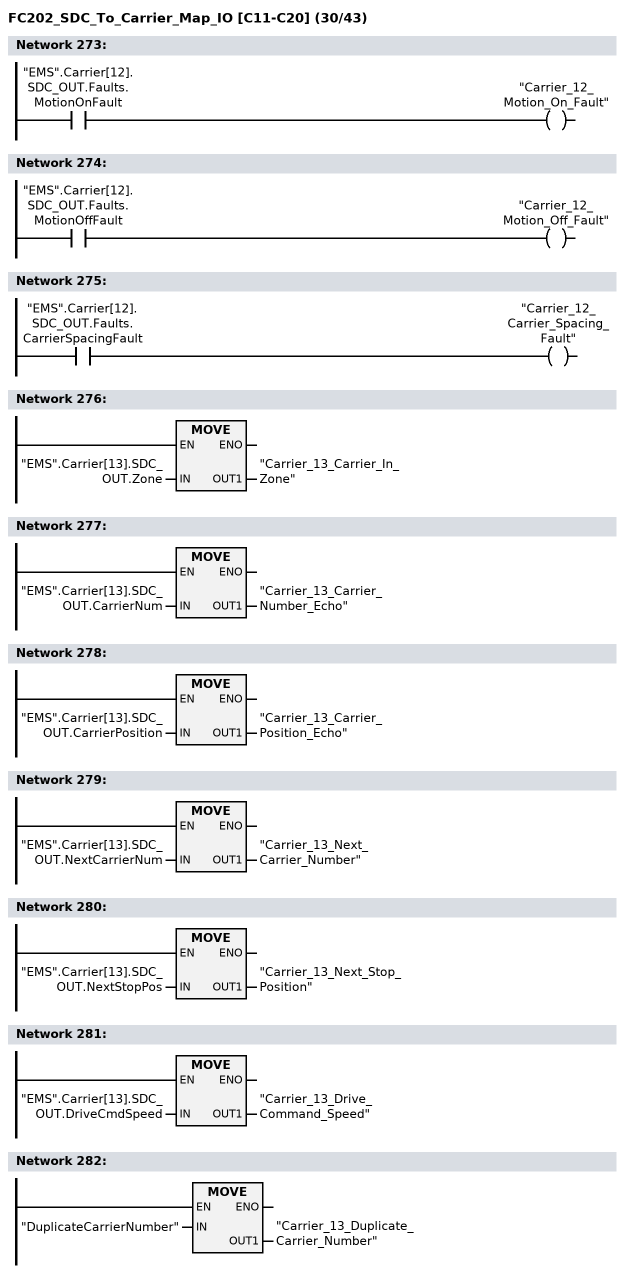
   RUNG wire#powerrail
      Contact( "EMS".Carrier[12].SDC_OUT.Faults.MotionOnFault )
      Coil( "Carrier_12_Motion_On_Fault" )
   END_RUNG
   // the same network as SCL:
   "Carrier_12_Motion_On_Fault" := "EMS".Carrier[12].SDC_OUT.Faults.MotionOnFault;
END_REGION

REGION Network 274
   RUNG wire#powerrail
      Contact( "EMS".Carrier[12].SDC_OUT.Faults.MotionOffFault )
      Coil( "Carrier_12_Motion_Off_Fault" )
   END_RUNG
   // the same network as SCL:
   "Carrier_12_Motion_Off_Fault" := "EMS".Carrier[12].SDC_OUT.Faults.MotionOffFault;
END_REGION

REGION Network 275
   RUNG wire#powerrail
      Contact( "EMS".Carrier[12].SDC_OUT.Faults.CarrierSpacingFault )
      Coil( "Carrier_12_Carrier_Spacing_Fault" )
   END_RUNG
   // the same network as SCL:
   "Carrier_12_Carrier_Spacing_Fault" := "EMS".Carrier[12].SDC_OUT.Faults.CarrierSpacingFault;
END_REGION

REGION Network 276
   RUNG wire#powerrail
      Move(in := "EMS".Carrier[13].SDC_OUT.Zone, out1 => "Carrier_13_Carrier_In_Zone")
   END_RUNG
   // the same network as SCL:
   "Carrier_13_Carrier_In_Zone" := "EMS".Carrier[13].SDC_OUT.Zone;
END_REGION

REGION Network 277
   RUNG wire#powerrail
      Move(in := "EMS".Carrier[13].SDC_OUT.CarrierNum, out1 => "Carrier_13_Carrier_Number_Echo")
   END_RUNG
   // the same network as SCL:
   "Carrier_13_Carrier_Number_Echo" := "EMS".Carrier[13].SDC_OUT.CarrierNum;
END_REGION

REGION Network 278
   RUNG wire#powerrail
      Move(in := "EMS".Carrier[13].SDC_OUT.CarrierPosition, out1 => "Carrier_13_Carrier_Position_Echo")
   END_RUNG
   // the same network as SCL:
   "Carrier_13_Carrier_Position_Echo" := "EMS".Carrier[13].SDC_OUT.CarrierPosition;
END_REGION

REGION Network 279
   RUNG wire#powerrail
      Move(in := "EMS".Carrier[13].SDC_OUT.NextCarrierNum, out1 => "Carrier_13_Next_Carrier_Number")
   END_RUNG
   // the same network as SCL:
   "Carrier_13_Next_Carrier_Number" := "EMS".Carrier[13].SDC_OUT.NextCarrierNum;
END_REGION

REGION Network 280
   RUNG wire#powerrail
      Move(in := "EMS".Carrier[13].SDC_OUT.NextStopPos, out1 => "Carrier_13_Next_Stop_Position")
   END_RUNG
   // the same network as SCL:
   "Carrier_13_Next_Stop_Position" := "EMS".Carrier[13].SDC_OUT.NextStopPos;
END_REGION

REGION Network 281
   RUNG wire#powerrail
      Move(in := "EMS".Carrier[13].SDC_OUT.DriveCmdSpeed, out1 => "Carrier_13_Drive_Command_Speed")
   END_RUNG
   // the same network as SCL:
   "Carrier_13_Drive_Command_Speed" := "EMS".Carrier[13].SDC_OUT.DriveCmdSpeed;
END_REGION

REGION Network 282
   RUNG wire#powerrail
      Move(in := "DuplicateCarrierNumber", out1 => "Carrier_13_Duplicate_Carrier_Number")
   END_RUNG
   // the same network as SCL:
   "Carrier_13_Duplicate_Carrier_Number" := "DuplicateCarrierNumber";
END_REGION

REGION Network 283
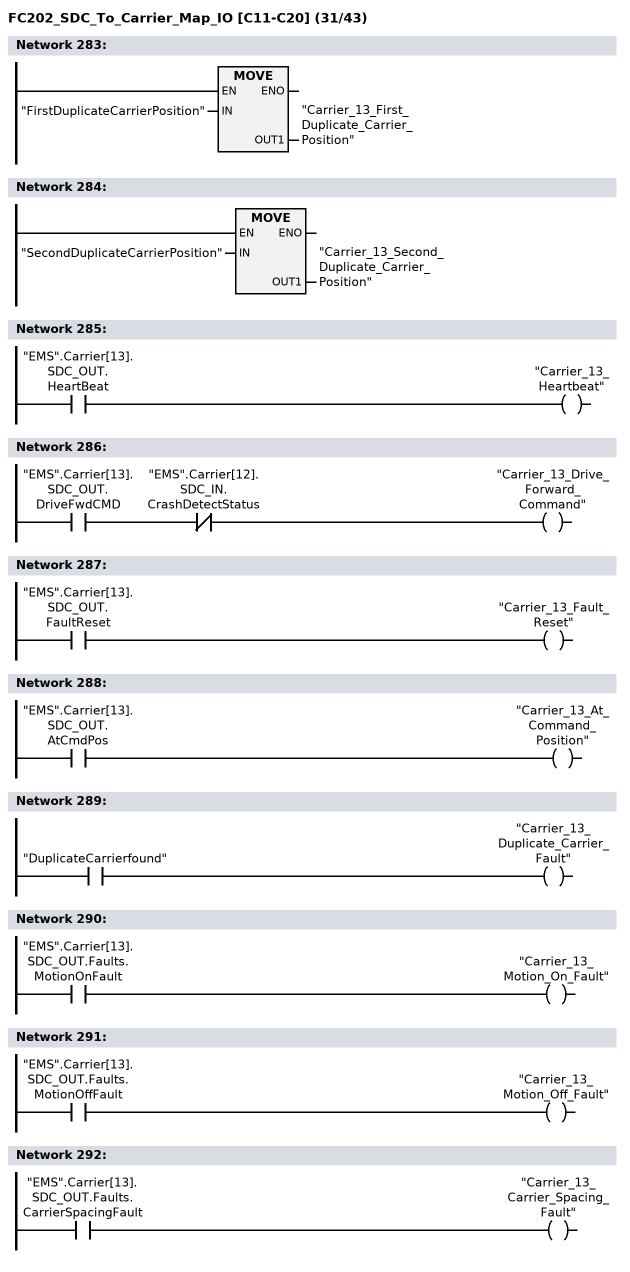
   RUNG wire#powerrail
      Move(in := "FirstDuplicateCarrierPosition", out1 => "Carrier_13_First_Duplicate_Carrier_Position")
   END_RUNG
   // the same network as SCL:
   "Carrier_13_First_Duplicate_Carrier_Position" := "FirstDuplicateCarrierPosition";
END_REGION

REGION Network 284
   RUNG wire#powerrail
      Move(in := "SecondDuplicateCarrierPosition", out1 => "Carrier_13_Second_Duplicate_Carrier_Position")
   END_RUNG
   // the same network as SCL:
   "Carrier_13_Second_Duplicate_Carrier_Position" := "SecondDuplicateCarrierPosition";
END_REGION

REGION Network 285
   RUNG wire#powerrail
      Contact( "EMS".Carrier[13].SDC_OUT.HeartBeat )
      Coil( "Carrier_13_Heartbeat" )
   END_RUNG
   // the same network as SCL:
   "Carrier_13_Heartbeat" := "EMS".Carrier[13].SDC_OUT.HeartBeat;
END_REGION

REGION Network 286
   RUNG wire#powerrail
      Contact( "EMS".Carrier[13].SDC_OUT.DriveFwdCMD )
      I_Contact( "EMS".Carrier[12].SDC_IN.CrashDetectStatus )
      Coil( "Carrier_13_Drive_Forward_Command" )
   END_RUNG
   // the same network as SCL:
   "Carrier_13_Drive_Forward_Command" := "EMS".Carrier[13].SDC_OUT.DriveFwdCMD AND NOT "EMS".Carrier[12].SDC_IN.CrashDetectStatus;
END_REGION

REGION Network 287
   RUNG wire#powerrail
      Contact( "EMS".Carrier[13].SDC_OUT.FaultReset )
      Coil( "Carrier_13_Fault_Reset" )
   END_RUNG
   // the same network as SCL:
   "Carrier_13_Fault_Reset" := "EMS".Carrier[13].SDC_OUT.FaultReset;
END_REGION

REGION Network 288
   RUNG wire#powerrail
      Contact( "EMS".Carrier[13].SDC_OUT.AtCmdPos )
      Coil( "Carrier_13_At_Command_Position" )
   END_RUNG
   // the same network as SCL:
   "Carrier_13_At_Command_Position" := "EMS".Carrier[13].SDC_OUT.AtCmdPos;
END_REGION

REGION Network 289
   RUNG wire#powerrail
      Contact( "DuplicateCarrierfound" )
      Coil( "Carrier_13_Duplicate_Carrier_Fault" )
   END_RUNG
   // the same network as SCL:
   "Carrier_13_Duplicate_Carrier_Fault" := "DuplicateCarrierfound";
END_REGION

REGION Network 290
   RUNG wire#powerrail
      Contact( "EMS".Carrier[13].SDC_OUT.Faults.MotionOnFault )
      Coil( "Carrier_13_Motion_On_Fault" )
   END_RUNG
   // the same network as SCL:
   "Carrier_13_Motion_On_Fault" := "EMS".Carrier[13].SDC_OUT.Faults.MotionOnFault;
END_REGION

REGION Network 291
   RUNG wire#powerrail
      Contact( "EMS".Carrier[13].SDC_OUT.Faults.MotionOffFault )
      Coil( "Carrier_13_Motion_Off_Fault" )
   END_RUNG
   // the same network as SCL:
   "Carrier_13_Motion_Off_Fault" := "EMS".Carrier[13].SDC_OUT.Faults.MotionOffFault;
END_REGION

REGION Network 292
   RUNG wire#powerrail
      Contact( "EMS".Carrier[13].SDC_OUT.Faults.CarrierSpacingFault )
      Coil( "Carrier_13_Carrier_Spacing_Fault" )
   END_RUNG
   // the same network as SCL:
   "Carrier_13_Carrier_Spacing_Fault" := "EMS".Carrier[13].SDC_OUT.Faults.CarrierSpacingFault;
END_REGION

REGION Network 293
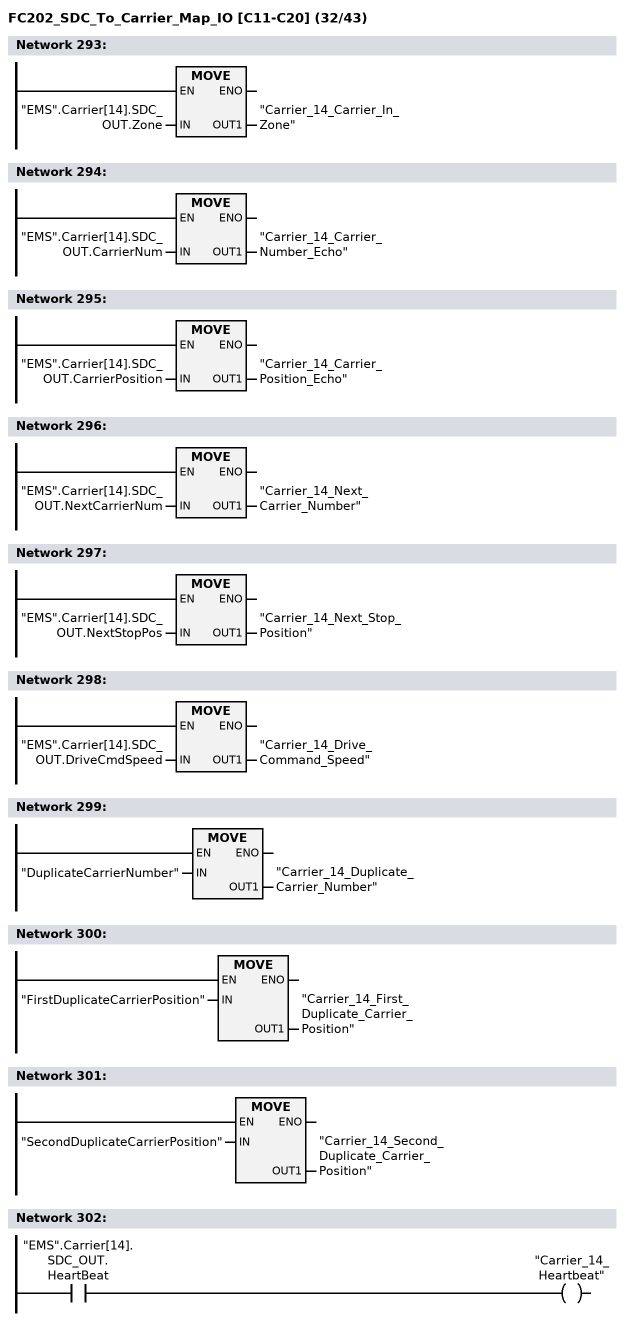
   RUNG wire#powerrail
      Move(in := "EMS".Carrier[14].SDC_OUT.Zone, out1 => "Carrier_14_Carrier_In_Zone")
   END_RUNG
   // the same network as SCL:
   "Carrier_14_Carrier_In_Zone" := "EMS".Carrier[14].SDC_OUT.Zone;
END_REGION

REGION Network 294
   RUNG wire#powerrail
      Move(in := "EMS".Carrier[14].SDC_OUT.CarrierNum, out1 => "Carrier_14_Carrier_Number_Echo")
   END_RUNG
   // the same network as SCL:
   "Carrier_14_Carrier_Number_Echo" := "EMS".Carrier[14].SDC_OUT.CarrierNum;
END_REGION

REGION Network 295
   RUNG wire#powerrail
      Move(in := "EMS".Carrier[14].SDC_OUT.CarrierPosition, out1 => "Carrier_14_Carrier_Position_Echo")
   END_RUNG
   // the same network as SCL:
   "Carrier_14_Carrier_Position_Echo" := "EMS".Carrier[14].SDC_OUT.CarrierPosition;
END_REGION

REGION Network 296
   RUNG wire#powerrail
      Move(in := "EMS".Carrier[14].SDC_OUT.NextCarrierNum, out1 => "Carrier_14_Next_Carrier_Number")
   END_RUNG
   // the same network as SCL:
   "Carrier_14_Next_Carrier_Number" := "EMS".Carrier[14].SDC_OUT.NextCarrierNum;
END_REGION

REGION Network 297
   RUNG wire#powerrail
      Move(in := "EMS".Carrier[14].SDC_OUT.NextStopPos, out1 => "Carrier_14_Next_Stop_Position")
   END_RUNG
   // the same network as SCL:
   "Carrier_14_Next_Stop_Position" := "EMS".Carrier[14].SDC_OUT.NextStopPos;
END_REGION

REGION Network 298
   RUNG wire#powerrail
      Move(in := "EMS".Carrier[14].SDC_OUT.DriveCmdSpeed, out1 => "Carrier_14_Drive_Command_Speed")
   END_RUNG
   // the same network as SCL:
   "Carrier_14_Drive_Command_Speed" := "EMS".Carrier[14].SDC_OUT.DriveCmdSpeed;
END_REGION

REGION Network 299
   RUNG wire#powerrail
      Move(in := "DuplicateCarrierNumber", out1 => "Carrier_14_Duplicate_Carrier_Number")
   END_RUNG
   // the same network as SCL:
   "Carrier_14_Duplicate_Carrier_Number" := "DuplicateCarrierNumber";
END_REGION

REGION Network 300
   RUNG wire#powerrail
      Move(in := "FirstDuplicateCarrierPosition", out1 => "Carrier_14_First_Duplicate_Carrier_Position")
   END_RUNG
   // the same network as SCL:
   "Carrier_14_First_Duplicate_Carrier_Position" := "FirstDuplicateCarrierPosition";
END_REGION

REGION Network 301
   RUNG wire#powerrail
      Move(in := "SecondDuplicateCarrierPosition", out1 => "Carrier_14_Second_Duplicate_Carrier_Position")
   END_RUNG
   // the same network as SCL:
   "Carrier_14_Second_Duplicate_Carrier_Position" := "SecondDuplicateCarrierPosition";
END_REGION

REGION Network 302
   RUNG wire#powerrail
      Contact( "EMS".Carrier[14].SDC_OUT.HeartBeat )
      Coil( "Carrier_14_Heartbeat" )
   END_RUNG
   // the same network as SCL:
   "Carrier_14_Heartbeat" := "EMS".Carrier[14].SDC_OUT.HeartBeat;
END_REGION

REGION Network 303
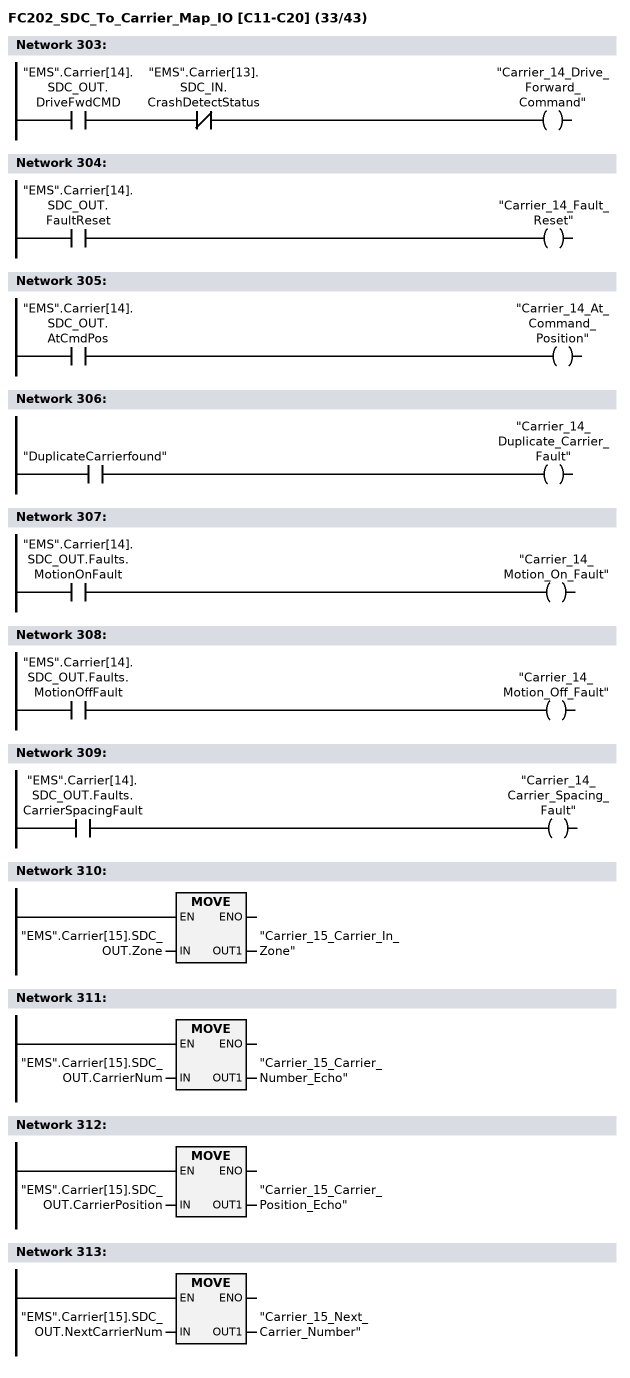
   RUNG wire#powerrail
      Contact( "EMS".Carrier[14].SDC_OUT.DriveFwdCMD )
      I_Contact( "EMS".Carrier[13].SDC_IN.CrashDetectStatus )
      Coil( "Carrier_14_Drive_Forward_Command" )
   END_RUNG
   // the same network as SCL:
   "Carrier_14_Drive_Forward_Command" := "EMS".Carrier[14].SDC_OUT.DriveFwdCMD AND NOT "EMS".Carrier[13].SDC_IN.CrashDetectStatus;
END_REGION

REGION Network 304
   RUNG wire#powerrail
      Contact( "EMS".Carrier[14].SDC_OUT.FaultReset )
      Coil( "Carrier_14_Fault_Reset" )
   END_RUNG
   // the same network as SCL:
   "Carrier_14_Fault_Reset" := "EMS".Carrier[14].SDC_OUT.FaultReset;
END_REGION

REGION Network 305
   RUNG wire#powerrail
      Contact( "EMS".Carrier[14].SDC_OUT.AtCmdPos )
      Coil( "Carrier_14_At_Command_Position" )
   END_RUNG
   // the same network as SCL:
   "Carrier_14_At_Command_Position" := "EMS".Carrier[14].SDC_OUT.AtCmdPos;
END_REGION

REGION Network 306
   RUNG wire#powerrail
      Contact( "DuplicateCarrierfound" )
      Coil( "Carrier_14_Duplicate_Carrier_Fault" )
   END_RUNG
   // the same network as SCL:
   "Carrier_14_Duplicate_Carrier_Fault" := "DuplicateCarrierfound";
END_REGION

REGION Network 307
   RUNG wire#powerrail
      Contact( "EMS".Carrier[14].SDC_OUT.Faults.MotionOnFault )
      Coil( "Carrier_14_Motion_On_Fault" )
   END_RUNG
   // the same network as SCL:
   "Carrier_14_Motion_On_Fault" := "EMS".Carrier[14].SDC_OUT.Faults.MotionOnFault;
END_REGION

REGION Network 308
   RUNG wire#powerrail
      Contact( "EMS".Carrier[14].SDC_OUT.Faults.MotionOffFault )
      Coil( "Carrier_14_Motion_Off_Fault" )
   END_RUNG
   // the same network as SCL:
   "Carrier_14_Motion_Off_Fault" := "EMS".Carrier[14].SDC_OUT.Faults.MotionOffFault;
END_REGION

REGION Network 309
   RUNG wire#powerrail
      Contact( "EMS".Carrier[14].SDC_OUT.Faults.CarrierSpacingFault )
      Coil( "Carrier_14_Carrier_Spacing_Fault" )
   END_RUNG
   // the same network as SCL:
   "Carrier_14_Carrier_Spacing_Fault" := "EMS".Carrier[14].SDC_OUT.Faults.CarrierSpacingFault;
END_REGION

REGION Network 310
   RUNG wire#powerrail
      Move(in := "EMS".Carrier[15].SDC_OUT.Zone, out1 => "Carrier_15_Carrier_In_Zone")
   END_RUNG
   // the same network as SCL:
   "Carrier_15_Carrier_In_Zone" := "EMS".Carrier[15].SDC_OUT.Zone;
END_REGION

REGION Network 311
   RUNG wire#powerrail
      Move(in := "EMS".Carrier[15].SDC_OUT.CarrierNum, out1 => "Carrier_15_Carrier_Number_Echo")
   END_RUNG
   // the same network as SCL:
   "Carrier_15_Carrier_Number_Echo" := "EMS".Carrier[15].SDC_OUT.CarrierNum;
END_REGION

REGION Network 312
   RUNG wire#powerrail
      Move(in := "EMS".Carrier[15].SDC_OUT.CarrierPosition, out1 => "Carrier_15_Carrier_Position_Echo")
   END_RUNG
   // the same network as SCL:
   "Carrier_15_Carrier_Position_Echo" := "EMS".Carrier[15].SDC_OUT.CarrierPosition;
END_REGION

REGION Network 313
   RUNG wire#powerrail
      Move(in := "EMS".Carrier[15].SDC_OUT.NextCarrierNum, out1 => "Carrier_15_Next_Carrier_Number")
   END_RUNG
   // the same network as SCL:
   "Carrier_15_Next_Carrier_Number" := "EMS".Carrier[15].SDC_OUT.NextCarrierNum;
END_REGION

REGION Network 314
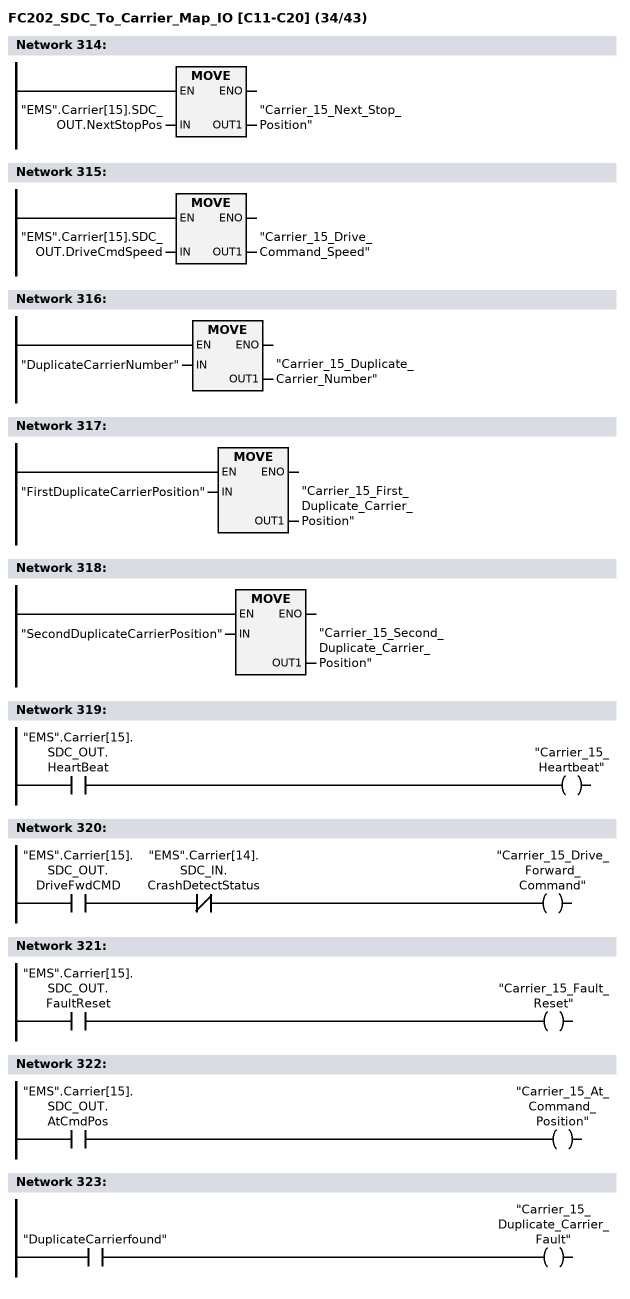
   RUNG wire#powerrail
      Move(in := "EMS".Carrier[15].SDC_OUT.NextStopPos, out1 => "Carrier_15_Next_Stop_Position")
   END_RUNG
   // the same network as SCL:
   "Carrier_15_Next_Stop_Position" := "EMS".Carrier[15].SDC_OUT.NextStopPos;
END_REGION

REGION Network 315
   RUNG wire#powerrail
      Move(in := "EMS".Carrier[15].SDC_OUT.DriveCmdSpeed, out1 => "Carrier_15_Drive_Command_Speed")
   END_RUNG
   // the same network as SCL:
   "Carrier_15_Drive_Command_Speed" := "EMS".Carrier[15].SDC_OUT.DriveCmdSpeed;
END_REGION

REGION Network 316
   RUNG wire#powerrail
      Move(in := "DuplicateCarrierNumber", out1 => "Carrier_15_Duplicate_Carrier_Number")
   END_RUNG
   // the same network as SCL:
   "Carrier_15_Duplicate_Carrier_Number" := "DuplicateCarrierNumber";
END_REGION

REGION Network 317
   RUNG wire#powerrail
      Move(in := "FirstDuplicateCarrierPosition", out1 => "Carrier_15_First_Duplicate_Carrier_Position")
   END_RUNG
   // the same network as SCL:
   "Carrier_15_First_Duplicate_Carrier_Position" := "FirstDuplicateCarrierPosition";
END_REGION

REGION Network 318
   RUNG wire#powerrail
      Move(in := "SecondDuplicateCarrierPosition", out1 => "Carrier_15_Second_Duplicate_Carrier_Position")
   END_RUNG
   // the same network as SCL:
   "Carrier_15_Second_Duplicate_Carrier_Position" := "SecondDuplicateCarrierPosition";
END_REGION

REGION Network 319
   RUNG wire#powerrail
      Contact( "EMS".Carrier[15].SDC_OUT.HeartBeat )
      Coil( "Carrier_15_Heartbeat" )
   END_RUNG
   // the same network as SCL:
   "Carrier_15_Heartbeat" := "EMS".Carrier[15].SDC_OUT.HeartBeat;
END_REGION

REGION Network 320
   RUNG wire#powerrail
      Contact( "EMS".Carrier[15].SDC_OUT.DriveFwdCMD )
      I_Contact( "EMS".Carrier[14].SDC_IN.CrashDetectStatus )
      Coil( "Carrier_15_Drive_Forward_Command" )
   END_RUNG
   // the same network as SCL:
   "Carrier_15_Drive_Forward_Command" := "EMS".Carrier[15].SDC_OUT.DriveFwdCMD AND NOT "EMS".Carrier[14].SDC_IN.CrashDetectStatus;
END_REGION

REGION Network 321
   RUNG wire#powerrail
      Contact( "EMS".Carrier[15].SDC_OUT.FaultReset )
      Coil( "Carrier_15_Fault_Reset" )
   END_RUNG
   // the same network as SCL:
   "Carrier_15_Fault_Reset" := "EMS".Carrier[15].SDC_OUT.FaultReset;
END_REGION

REGION Network 322
   RUNG wire#powerrail
      Contact( "EMS".Carrier[15].SDC_OUT.AtCmdPos )
      Coil( "Carrier_15_At_Command_Position" )
   END_RUNG
   // the same network as SCL:
   "Carrier_15_At_Command_Position" := "EMS".Carrier[15].SDC_OUT.AtCmdPos;
END_REGION

REGION Network 323
   RUNG wire#powerrail
      Contact( "DuplicateCarrierfound" )
      Coil( "Carrier_15_Duplicate_Carrier_Fault" )
   END_RUNG
   // the same network as SCL:
   "Carrier_15_Duplicate_Carrier_Fault" := "DuplicateCarrierfound";
END_REGION

REGION Network 324
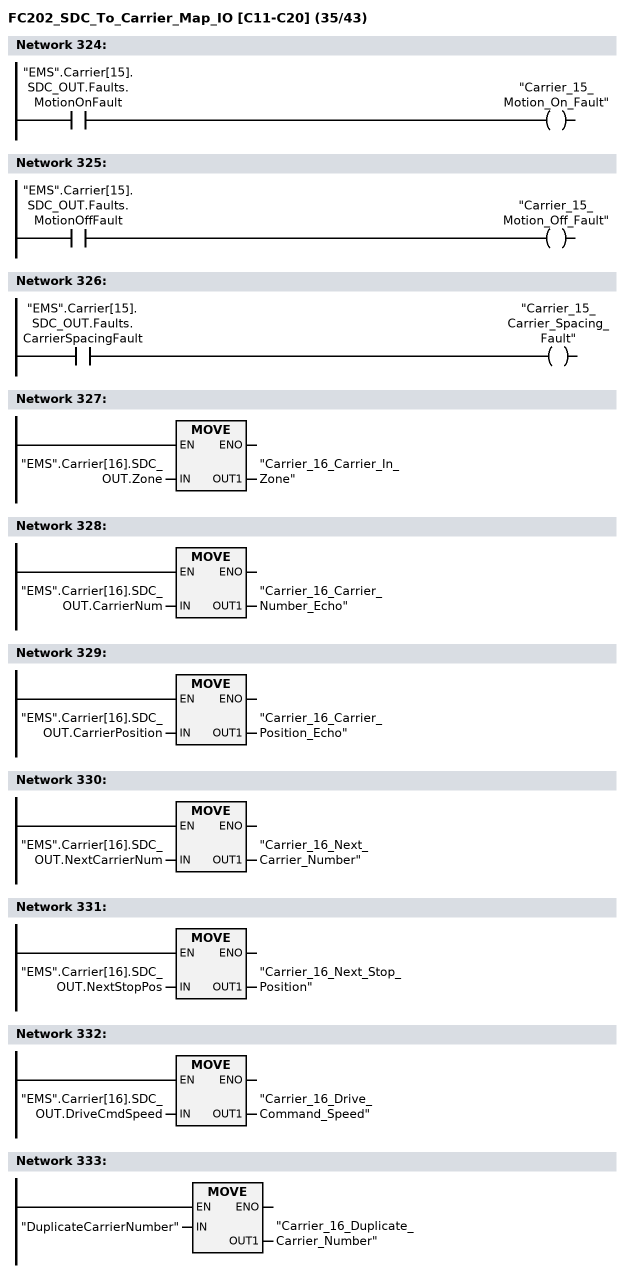
   RUNG wire#powerrail
      Contact( "EMS".Carrier[15].SDC_OUT.Faults.MotionOnFault )
      Coil( "Carrier_15_Motion_On_Fault" )
   END_RUNG
   // the same network as SCL:
   "Carrier_15_Motion_On_Fault" := "EMS".Carrier[15].SDC_OUT.Faults.MotionOnFault;
END_REGION

REGION Network 325
   RUNG wire#powerrail
      Contact( "EMS".Carrier[15].SDC_OUT.Faults.MotionOffFault )
      Coil( "Carrier_15_Motion_Off_Fault" )
   END_RUNG
   // the same network as SCL:
   "Carrier_15_Motion_Off_Fault" := "EMS".Carrier[15].SDC_OUT.Faults.MotionOffFault;
END_REGION

REGION Network 326
   RUNG wire#powerrail
      Contact( "EMS".Carrier[15].SDC_OUT.Faults.CarrierSpacingFault )
      Coil( "Carrier_15_Carrier_Spacing_Fault" )
   END_RUNG
   // the same network as SCL:
   "Carrier_15_Carrier_Spacing_Fault" := "EMS".Carrier[15].SDC_OUT.Faults.CarrierSpacingFault;
END_REGION

REGION Network 327
   RUNG wire#powerrail
      Move(in := "EMS".Carrier[16].SDC_OUT.Zone, out1 => "Carrier_16_Carrier_In_Zone")
   END_RUNG
   // the same network as SCL:
   "Carrier_16_Carrier_In_Zone" := "EMS".Carrier[16].SDC_OUT.Zone;
END_REGION

REGION Network 328
   RUNG wire#powerrail
      Move(in := "EMS".Carrier[16].SDC_OUT.CarrierNum, out1 => "Carrier_16_Carrier_Number_Echo")
   END_RUNG
   // the same network as SCL:
   "Carrier_16_Carrier_Number_Echo" := "EMS".Carrier[16].SDC_OUT.CarrierNum;
END_REGION

REGION Network 329
   RUNG wire#powerrail
      Move(in := "EMS".Carrier[16].SDC_OUT.CarrierPosition, out1 => "Carrier_16_Carrier_Position_Echo")
   END_RUNG
   // the same network as SCL:
   "Carrier_16_Carrier_Position_Echo" := "EMS".Carrier[16].SDC_OUT.CarrierPosition;
END_REGION

REGION Network 330
   RUNG wire#powerrail
      Move(in := "EMS".Carrier[16].SDC_OUT.NextCarrierNum, out1 => "Carrier_16_Next_Carrier_Number")
   END_RUNG
   // the same network as SCL:
   "Carrier_16_Next_Carrier_Number" := "EMS".Carrier[16].SDC_OUT.NextCarrierNum;
END_REGION

REGION Network 331
   RUNG wire#powerrail
      Move(in := "EMS".Carrier[16].SDC_OUT.NextStopPos, out1 => "Carrier_16_Next_Stop_Position")
   END_RUNG
   // the same network as SCL:
   "Carrier_16_Next_Stop_Position" := "EMS".Carrier[16].SDC_OUT.NextStopPos;
END_REGION

REGION Network 332
   RUNG wire#powerrail
      Move(in := "EMS".Carrier[16].SDC_OUT.DriveCmdSpeed, out1 => "Carrier_16_Drive_Command_Speed")
   END_RUNG
   // the same network as SCL:
   "Carrier_16_Drive_Command_Speed" := "EMS".Carrier[16].SDC_OUT.DriveCmdSpeed;
END_REGION

REGION Network 333
   RUNG wire#powerrail
      Move(in := "DuplicateCarrierNumber", out1 => "Carrier_16_Duplicate_Carrier_Number")
   END_RUNG
   // the same network as SCL:
   "Carrier_16_Duplicate_Carrier_Number" := "DuplicateCarrierNumber";
END_REGION

REGION Network 334
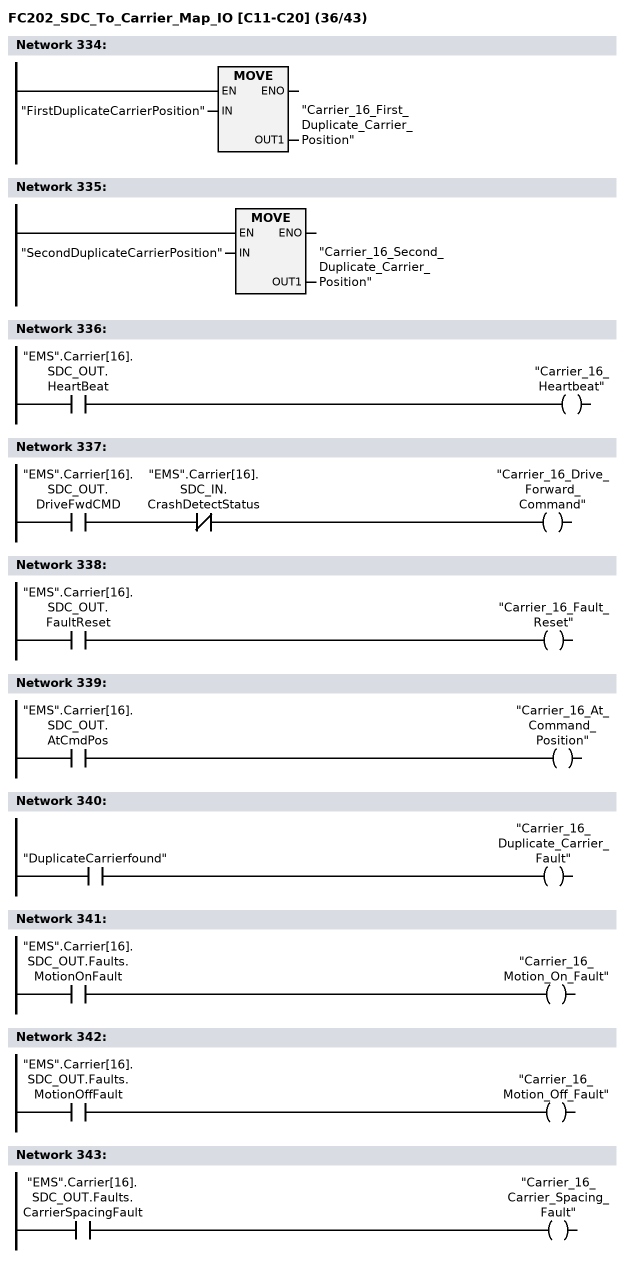
   RUNG wire#powerrail
      Move(in := "FirstDuplicateCarrierPosition", out1 => "Carrier_16_First_Duplicate_Carrier_Position")
   END_RUNG
   // the same network as SCL:
   "Carrier_16_First_Duplicate_Carrier_Position" := "FirstDuplicateCarrierPosition";
END_REGION

REGION Network 335
   RUNG wire#powerrail
      Move(in := "SecondDuplicateCarrierPosition", out1 => "Carrier_16_Second_Duplicate_Carrier_Position")
   END_RUNG
   // the same network as SCL:
   "Carrier_16_Second_Duplicate_Carrier_Position" := "SecondDuplicateCarrierPosition";
END_REGION

REGION Network 336
   RUNG wire#powerrail
      Contact( "EMS".Carrier[16].SDC_OUT.HeartBeat )
      Coil( "Carrier_16_Heartbeat" )
   END_RUNG
   // the same network as SCL:
   "Carrier_16_Heartbeat" := "EMS".Carrier[16].SDC_OUT.HeartBeat;
END_REGION

REGION Network 337
   RUNG wire#powerrail
      Contact( "EMS".Carrier[16].SDC_OUT.DriveFwdCMD )
      I_Contact( "EMS".Carrier[16].SDC_IN.CrashDetectStatus )
      Coil( "Carrier_16_Drive_Forward_Command" )
   END_RUNG
   // the same network as SCL:
   "Carrier_16_Drive_Forward_Command" := "EMS".Carrier[16].SDC_OUT.DriveFwdCMD AND NOT "EMS".Carrier[16].SDC_IN.CrashDetectStatus;
END_REGION

REGION Network 338
   RUNG wire#powerrail
      Contact( "EMS".Carrier[16].SDC_OUT.FaultReset )
      Coil( "Carrier_16_Fault_Reset" )
   END_RUNG
   // the same network as SCL:
   "Carrier_16_Fault_Reset" := "EMS".Carrier[16].SDC_OUT.FaultReset;
END_REGION

REGION Network 339
   RUNG wire#powerrail
      Contact( "EMS".Carrier[16].SDC_OUT.AtCmdPos )
      Coil( "Carrier_16_At_Command_Position" )
   END_RUNG
   // the same network as SCL:
   "Carrier_16_At_Command_Position" := "EMS".Carrier[16].SDC_OUT.AtCmdPos;
END_REGION

REGION Network 340
   RUNG wire#powerrail
      Contact( "DuplicateCarrierfound" )
      Coil( "Carrier_16_Duplicate_Carrier_Fault" )
   END_RUNG
   // the same network as SCL:
   "Carrier_16_Duplicate_Carrier_Fault" := "DuplicateCarrierfound";
END_REGION

REGION Network 341
   RUNG wire#powerrail
      Contact( "EMS".Carrier[16].SDC_OUT.Faults.MotionOnFault )
      Coil( "Carrier_16_Motion_On_Fault" )
   END_RUNG
   // the same network as SCL:
   "Carrier_16_Motion_On_Fault" := "EMS".Carrier[16].SDC_OUT.Faults.MotionOnFault;
END_REGION

REGION Network 342
   RUNG wire#powerrail
      Contact( "EMS".Carrier[16].SDC_OUT.Faults.MotionOffFault )
      Coil( "Carrier_16_Motion_Off_Fault" )
   END_RUNG
   // the same network as SCL:
   "Carrier_16_Motion_Off_Fault" := "EMS".Carrier[16].SDC_OUT.Faults.MotionOffFault;
END_REGION

REGION Network 343
   RUNG wire#powerrail
      Contact( "EMS".Carrier[16].SDC_OUT.Faults.CarrierSpacingFault )
      Coil( "Carrier_16_Carrier_Spacing_Fault" )
   END_RUNG
   // the same network as SCL:
   "Carrier_16_Carrier_Spacing_Fault" := "EMS".Carrier[16].SDC_OUT.Faults.CarrierSpacingFault;
END_REGION

REGION Network 344
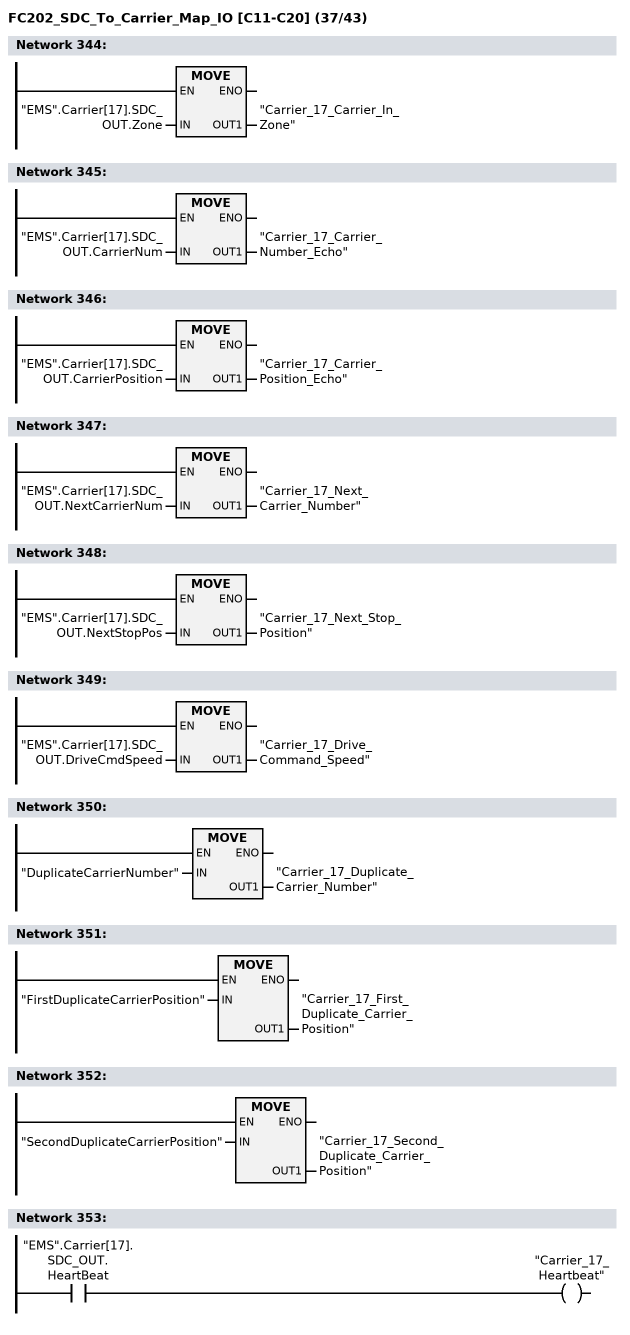
   RUNG wire#powerrail
      Move(in := "EMS".Carrier[17].SDC_OUT.Zone, out1 => "Carrier_17_Carrier_In_Zone")
   END_RUNG
   // the same network as SCL:
   "Carrier_17_Carrier_In_Zone" := "EMS".Carrier[17].SDC_OUT.Zone;
END_REGION

REGION Network 345
   RUNG wire#powerrail
      Move(in := "EMS".Carrier[17].SDC_OUT.CarrierNum, out1 => "Carrier_17_Carrier_Number_Echo")
   END_RUNG
   // the same network as SCL:
   "Carrier_17_Carrier_Number_Echo" := "EMS".Carrier[17].SDC_OUT.CarrierNum;
END_REGION

REGION Network 346
   RUNG wire#powerrail
      Move(in := "EMS".Carrier[17].SDC_OUT.CarrierPosition, out1 => "Carrier_17_Carrier_Position_Echo")
   END_RUNG
   // the same network as SCL:
   "Carrier_17_Carrier_Position_Echo" := "EMS".Carrier[17].SDC_OUT.CarrierPosition;
END_REGION

REGION Network 347
   RUNG wire#powerrail
      Move(in := "EMS".Carrier[17].SDC_OUT.NextCarrierNum, out1 => "Carrier_17_Next_Carrier_Number")
   END_RUNG
   // the same network as SCL:
   "Carrier_17_Next_Carrier_Number" := "EMS".Carrier[17].SDC_OUT.NextCarrierNum;
END_REGION

REGION Network 348
   RUNG wire#powerrail
      Move(in := "EMS".Carrier[17].SDC_OUT.NextStopPos, out1 => "Carrier_17_Next_Stop_Position")
   END_RUNG
   // the same network as SCL:
   "Carrier_17_Next_Stop_Position" := "EMS".Carrier[17].SDC_OUT.NextStopPos;
END_REGION

REGION Network 349
   RUNG wire#powerrail
      Move(in := "EMS".Carrier[17].SDC_OUT.DriveCmdSpeed, out1 => "Carrier_17_Drive_Command_Speed")
   END_RUNG
   // the same network as SCL:
   "Carrier_17_Drive_Command_Speed" := "EMS".Carrier[17].SDC_OUT.DriveCmdSpeed;
END_REGION

REGION Network 350
   RUNG wire#powerrail
      Move(in := "DuplicateCarrierNumber", out1 => "Carrier_17_Duplicate_Carrier_Number")
   END_RUNG
   // the same network as SCL:
   "Carrier_17_Duplicate_Carrier_Number" := "DuplicateCarrierNumber";
END_REGION

REGION Network 351
   RUNG wire#powerrail
      Move(in := "FirstDuplicateCarrierPosition", out1 => "Carrier_17_First_Duplicate_Carrier_Position")
   END_RUNG
   // the same network as SCL:
   "Carrier_17_First_Duplicate_Carrier_Position" := "FirstDuplicateCarrierPosition";
END_REGION

REGION Network 352
   RUNG wire#powerrail
      Move(in := "SecondDuplicateCarrierPosition", out1 => "Carrier_17_Second_Duplicate_Carrier_Position")
   END_RUNG
   // the same network as SCL:
   "Carrier_17_Second_Duplicate_Carrier_Position" := "SecondDuplicateCarrierPosition";
END_REGION

REGION Network 353
   RUNG wire#powerrail
      Contact( "EMS".Carrier[17].SDC_OUT.HeartBeat )
      Coil( "Carrier_17_Heartbeat" )
   END_RUNG
   // the same network as SCL:
   "Carrier_17_Heartbeat" := "EMS".Carrier[17].SDC_OUT.HeartBeat;
END_REGION

REGION Network 354
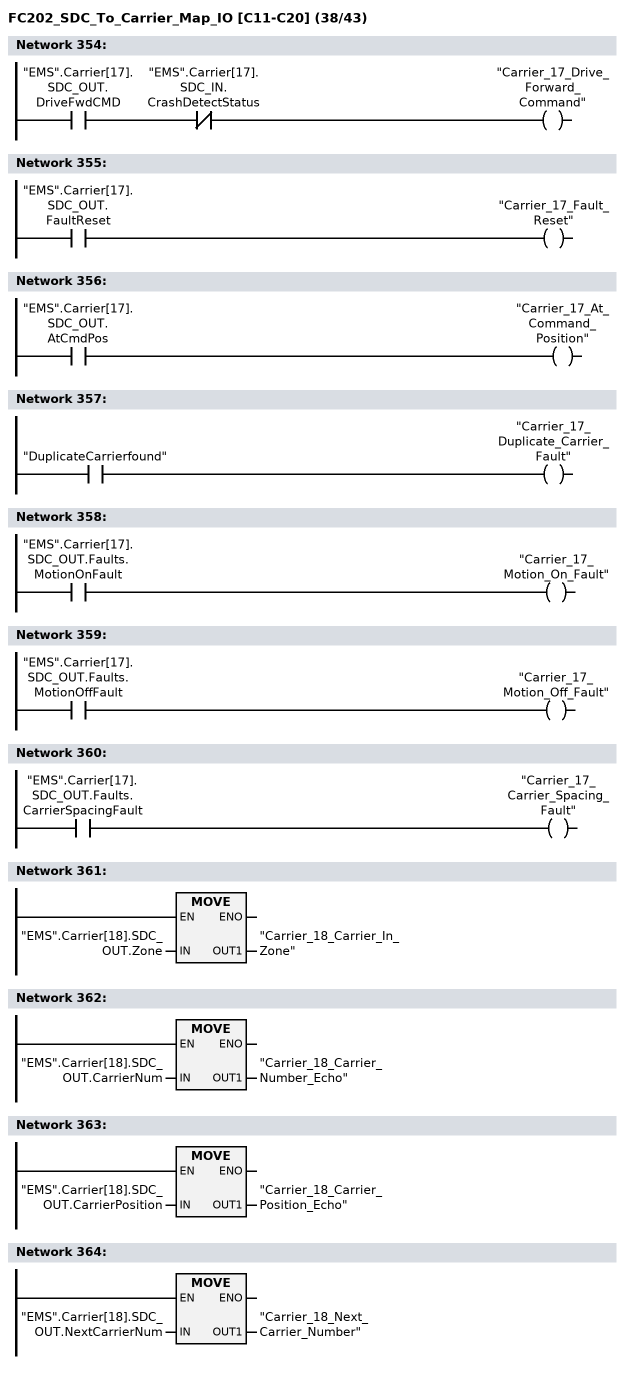
   RUNG wire#powerrail
      Contact( "EMS".Carrier[17].SDC_OUT.DriveFwdCMD )
      I_Contact( "EMS".Carrier[17].SDC_IN.CrashDetectStatus )
      Coil( "Carrier_17_Drive_Forward_Command" )
   END_RUNG
   // the same network as SCL:
   "Carrier_17_Drive_Forward_Command" := "EMS".Carrier[17].SDC_OUT.DriveFwdCMD AND NOT "EMS".Carrier[17].SDC_IN.CrashDetectStatus;
END_REGION

REGION Network 355
   RUNG wire#powerrail
      Contact( "EMS".Carrier[17].SDC_OUT.FaultReset )
      Coil( "Carrier_17_Fault_Reset" )
   END_RUNG
   // the same network as SCL:
   "Carrier_17_Fault_Reset" := "EMS".Carrier[17].SDC_OUT.FaultReset;
END_REGION

REGION Network 356
   RUNG wire#powerrail
      Contact( "EMS".Carrier[17].SDC_OUT.AtCmdPos )
      Coil( "Carrier_17_At_Command_Position" )
   END_RUNG
   // the same network as SCL:
   "Carrier_17_At_Command_Position" := "EMS".Carrier[17].SDC_OUT.AtCmdPos;
END_REGION
